
       // If a status for the inerting system changed by operator copy this to the select number and do not read all status values
       IF "DB614_MH_State".InertingMH["DB614_MH_State".ReadDeviceNo].Inert_ON_OFF <> "DB614_MH_State".InertingMH[0].Inert_ON_OFF OR
           "DB614_MH_State".InertingMH["DB614_MH_State".ReadDeviceNo].Enable_Purge <> "DB614_MH_State".InertingMH[0].Enable_Purge
       THEN
           "DB614_MH_State".InertingMH["DB614_MH_State".ReadDeviceNo].Inert_ON_OFF := "DB614_MH_State".InertingMH[0].Inert_ON_OFF;
           "DB614_MH_State".InertingMH["DB614_MH_State".ReadDeviceNo].Enable_Purge := "DB614_MH_State".InertingMH[0].Enable_Purge;
       ELSE
           "DB614_MH_State".InertingMH[0] := "DB614_MH_State".InertingMH["DB614_MH_State".ReadDeviceNo];
       END_IF;

   END_IF;

   // Copy the Status bits after changing
   IF "DB614_MH_State".Write THEN

       "DB614_MH_State".Write := False;

   END_IF;

   // Copy the values if nessesary
   IF "DB704_MH_Value".Write THEN
       "DB604_PV_Mixinghead".Mixinghead["DB614_MH_State".ReadDeviceNo] := "DB604_PV_Mixinghead".Mixinghead[0];
       "DB704_MH_Value".Mixinghead["DB614_MH_State".ReadDeviceNo] := "DB704_MH_Value".Mixinghead[0];
       "DB704_MH_Value".MH_Inerting["DB614_MH_State".ReadDeviceNo] := "DB704_MH_Value".MH_Inerting[0];

       "DB704_MH_Value".Write := False;

   END_IF;

   // Show the actual values every time:
   // 
   "DB604_PV_Mixinghead".Mixinghead[0].Pressure_Connection[1].PV_ActV := "DB604_PV_Mixinghead".Mixinghead["DB614_MH_State".ReadDeviceNo].Pressure_Connection[1].PV_ActV;
   "DB604_PV_Mixinghead".Mixinghead[0].Pressure_Connection[2].PV_ActV := "DB604_PV_Mixinghead".Mixinghead["DB614_MH_State".ReadDeviceNo].Pressure_Connection[2].PV_ActV;
   "DB604_PV_Mixinghead".Mixinghead[0].Pressure_Connection[3].PV_ActV := "DB604_PV_Mixinghead".Mixinghead["DB614_MH_State".ReadDeviceNo].Pressure_Connection[3].PV_ActV;
   "DB604_PV_Mixinghead".Mixinghead[0].Pressure_Connection[4].PV_ActV := "DB604_PV_Mixinghead".Mixinghead["DB614_MH_State".ReadDeviceNo].Pressure_Connection[4].PV_ActV;
   "DB604_PV_Mixinghead".Mixinghead[0].Pressure_Connection[5].PV_ActV := "DB604_PV_Mixinghead".Mixinghead["DB614_MH_State".ReadDeviceNo].Pressure_Connection[5].PV_ActV;
   "DB604_PV_Mixinghead".Mixinghead[0].Pressure_Connection[6].PV_ActV := "DB604_PV_Mixinghead".Mixinghead["DB614_MH_State".ReadDeviceNo].Pressure_Connection[6].PV_ActV;

   "DB604_PV_Mixinghead".Mixinghead[0].Temperature_Connection[1].PV_ActV := "DB604_PV_Mixinghead".Mixinghead["DB614_MH_State".ReadDeviceNo].Temperature_Connection[1].PV_ActV;
   "DB604_PV_Mixinghead".Mixinghead[0].Temperature_Connection[2].PV_ActV := "DB604_PV_Mixinghead".Mixinghead["DB614_MH_State".ReadDeviceNo].Temperature_Connection[2].PV_ActV;
   "DB604_PV_Mixinghead".Mixinghead[0].Temperature_Connection[3].PV_ActV := "DB604_PV_Mixinghead".Mixinghead["DB614_MH_State".ReadDeviceNo].Temperature_Connection[3].PV_ActV;
   "DB604_PV_Mixinghead".Mixinghead[0].Temperature_Connection[4].PV_ActV := "DB604_PV_Mixinghead".Mixinghead["DB614_MH_State".ReadDeviceNo].Temperature_Connection[4].PV_ActV;
   "DB604_PV_Mixinghead".Mixinghead[0].Temperature_Connection[5].PV_ActV := "DB604_PV_Mixinghead".Mixinghead["DB614_MH_State".ReadDeviceNo].Temperature_Connection[5].PV_ActV;
   "DB604_PV_Mixinghead".Mixinghead[0].Temperature_Connection[6].PV_ActV := "DB604_PV_Mixinghead".Mixinghead["DB614_MH_State".ReadDeviceNo].Temperature_Connection[6].PV_ActV;

   "DB604_PV_Mixinghead".Mixinghead[0].SteeringPiston.PV_ActV := "DB604_PV_Mixinghead".Mixinghead["DB614_MH_State".ReadDeviceNo].SteeringPiston.PV_ActV;
   "DB604_PV_Mixinghead".Mixinghead[0].CleaningPiston.PV_ActV := "DB604_PV_Mixinghead".Mixinghead["DB614_MH_State".ReadDeviceNo].CleaningPiston.PV_ActV;
   "DB604_PV_Mixinghead".Mixinghead[0].Inerting.PV_ActV := "DB604_PV_Mixinghead".Mixinghead["DB614_MH_State".ReadDeviceNo].Inerting.PV_ActV;

   // Show the in/ output from MH every time
   "DB123_MH_IO_Signals".MH[0] := "DB123_MH_IO_Signals".MH["DB614_MH_State".ReadDeviceNo];

   // Show the actual information about the selected mixinghead
   "DB614_MH_State".MH_Connection[0] := "DB614_MH_State".MH_Connection["DB614_MH_State".ReadDeviceNo];

   // Information about shot adjustment
   "DB614_MH_State".ShotAdjustMH[0] := "DB614_MH_State".ShotAdjustMH["DB614_MH_State".ReadDeviceNo];
END_FUNCTION

FUNCTION "FC5019_InterfaceInterface" : Void   // FC5019, SCL
{ S7_Optimized_Access := 'FALSE' }
VERSION : 0.1
   VAR_INPUT
      Enable : Bool;
   END_VAR
BEGIN
   // Status: DB612_Hydraulic_State
   // Read all status bits during window is selected and NO button is pressed
     IF "DB119_Interface_Visu".Read THEN
       "DB119_Interface_Visu".MouldCarrer[0] := "DB119_Interface_Visu".MouldCarrer["DB119_Interface_Visu".ReadWriteDeviceNo];
       "DB119_Interface_Visu".APInterface[0] := "DB119_Interface_Visu".APInterface["DB119_Interface_Visu".ReadWriteDeviceNo];
     END_IF;
END_FUNCTION

FUNCTION "FC5020_InterfaceConfig" : Void   // FC5020, SCL
{ S7_Optimized_Access := 'FALSE' }
VERSION : 0.1
   VAR_INPUT
      Enable : Bool;
   END_VAR
BEGIN

   // Values:  "DB1200_ProCanConf" 
     IF "DB1200_ProCanConf".Read OR "DB1200_ProCanConf".Write OR "DB1200_ProCanConf".Copy THEN
       IF "DB1200_ProCanConf".Read THEN
         "DB1200_ProCanConf".ProCanConf[0] := "DB1200_ProCanConf".ProCanConf["DB1200_ProCanConf".ReadWriteDeviceNo];
         "DB1200_ProCanConf".Read := FALSE;
       END_IF;
       IF "DB1200_ProCanConf".Write THEN
         "DB1200_ProCanConf".ProCanConf["DB1200_ProCanConf".ReadWriteDeviceNo] := "DB1200_ProCanConf".ProCanConf[0];
         "DB1200_ProCanConf".Write := FALSE;
       END_IF;
         IF "DB1200_ProCanConf".CopyDeviceNO >0 THEN
         IF "DB1200_ProCanConf".Copy THEN
             "DB1200_ProCanConf".ProCanConf["DB1200_ProCanConf".CopyDeviceNO] := "DB1200_ProCanConf".ProCanConf[0];
             "DB1200_ProCanConf".Copy := FALSE;
             "DB1200_ProCanConf".CopyDeviceNO := 0;
         END_IF;
        END_IF;
      END_IF;    

   // Values:  "DB1232_ProCanIO_MH" 
     IF "DB1232_ProCanIO_MH".Read OR "DB1232_ProCanIO_MH".Write OR "DB1232_ProCanIO_MH".Copy THEN
       IF "DB1232_ProCanIO_MH".Read THEN
         "DB1232_ProCanIO_MH".AddressMH[0] := "DB1232_ProCanIO_MH".AddressMH["DB1232_ProCanIO_MH".ReadWriteDeviceNo];
         "DB1232_ProCanIO_MH".Read := FALSE;
       END_IF;
       IF "DB1232_ProCanIO_MH".Write THEN
         "DB1232_ProCanIO_MH".AddressMH["DB1232_ProCanIO_MH".ReadWriteDeviceNo] := "DB1232_ProCanIO_MH".AddressMH[0];
         "DB1232_ProCanIO_MH".Write := FALSE;
       END_IF;
         IF "DB1232_ProCanIO_MH".CopyDeviceNO >0 THEN
         IF "DB1232_ProCanIO_MH".Copy THEN
             "DB1232_ProCanIO_MH".AddressMH["DB1232_ProCanIO_MH".CopyDeviceNO] := "DB1232_ProCanIO_MH".AddressMH[0];
             "DB1232_ProCanIO_MH".Copy := FALSE;
             "DB1232_ProCanIO_MH".CopyDeviceNO := 0;
         END_IF;
        END_IF;
      END_IF;

   // Values:  "DB1233_ProCanIO_Flow" 
     IF "DB1233_ProCanIO_Flow".Read OR "DB1233_ProCanIO_Flow".Write OR "DB1233_ProCanIO_Flow".Copy THEN
       IF "DB1233_ProCanIO_Flow".Read THEN
         "DB1233_ProCanIO_Flow".AddressFlow[0] := "DB1233_ProCanIO_Flow".AddressFlow["DB1233_ProCanIO_Flow".ReadWriteDeviceNo];
         "DB1233_ProCanIO_Flow".Read := FALSE;
       END_IF;
       IF "DB1233_ProCanIO_Flow".Write THEN
         "DB1233_ProCanIO_Flow".AddressFlow["DB1233_ProCanIO_Flow".ReadWriteDeviceNo] := "DB1233_ProCanIO_Flow".AddressFlow[0];
         "DB1233_ProCanIO_Flow".Write := FALSE;
       END_IF;
         IF "DB1233_ProCanIO_Flow".CopyDeviceNO >0 THEN
         IF "DB1233_ProCanIO_Flow".Copy THEN
             "DB1233_ProCanIO_Flow".AddressFlow["DB1233_ProCanIO_Flow".CopyDeviceNO] := "DB1233_ProCanIO_Flow".AddressFlow[0];
             "DB1233_ProCanIO_Flow".Copy := FALSE;
             "DB1233_ProCanIO_Flow".CopyDeviceNO := 0;
         END_IF;
        END_IF;
      END_IF;
END_FUNCTION

FUNCTION "FC5030_InterfaceactualMHValue" : Void   // FC5030, SCL
{ S7_Optimized_Access := 'FALSE' }
VERSION : 0.1
   VAR_INPUT
      IN_MachineNo : Int;
   END_VAR
   VAR_TEMP
      N : Int;
      i : Int;
      AmountComponent : Int;
      Temp_MachineNo : Byte;
   END_VAR
BEGIN
   // Baustein zur Ermittlung der akteullen Mischkopf- Informationen
   // 
   // 1. Maschine ist im Ruhestand, Kein Kreislauf oder Zyxklus aktiv
   //    Die Werte des zuerst freigegebenen Mischkopfes an dieser Maschine werden angezeigt
   //  
   #Temp_MachineNo := INT_TO_BYTE(#IN_MachineNo);
   //  
   "DB619_State_MPart".ActMHInerting[#IN_MachineNo].Total_Flow_N2_Visu := "DB614_MH_State".InertingMH[1].Total_Flow_N2_Visu;

   IF NOT "DB619_State_MPart".Recirculation[#IN_MachineNo].Is_active AND
      NOT "DB619_State_MPart".Cycle[#IN_MachineNo].running THEN

      "DB619_State_MPart".ActMHComponent[1].OP_Manual := 0;
      "DB619_State_MPart".ActMHComponent[1].OP_Automatic := 0;
      "DB619_State_MPart".ActMHComponent[1].OP_Service := 0;

     FOR #N := 1 TO "DB790_PlantParameter".AmountMH DO

       IF "DB704_MH_Value".Mixinghead[#N].MH_Active AND
           "DB704_MH_Value".Mixinghead[#N].MachineNumber = #Temp_MachineNo THEN

         "DB619_State_MPart".ActMHPressureMa[#IN_MachineNo].Comp[1] :=  "DB604_PV_Mixinghead".Mixinghead[#N].Pressure_Connection[1].PV_ActV.Value;
         "DB619_State_MPart".ActMHPressureMa[#IN_MachineNo].Comp[2] :=  "DB604_PV_Mixinghead".Mixinghead[#N].Pressure_Connection[2].PV_ActV.Value;
         "DB619_State_MPart".ActMHPressureMa[#IN_MachineNo].Comp[3] :=  "DB604_PV_Mixinghead".Mixinghead[#N].Pressure_Connection[3].PV_ActV.Value;
         "DB619_State_MPart".ActMHPressureMa[#IN_MachineNo].Comp[4] :=  "DB604_PV_Mixinghead".Mixinghead[#N].Pressure_Connection[4].PV_ActV.Value;
         "DB619_State_MPart".ActMHPressureMa[#IN_MachineNo].Comp[5] :=  "DB604_PV_Mixinghead".Mixinghead[#N].Pressure_Connection[5].PV_ActV.Value;
         "DB619_State_MPart".ActMHPressureMa[#IN_MachineNo].Comp[6] :=  "DB604_PV_Mixinghead".Mixinghead[#N].Pressure_Connection[6].PV_ActV.Value;
         "DB619_State_MPart".ActMHTemperatureMa[#IN_MachineNo].Comp[1] :=  "DB604_PV_Mixinghead".Mixinghead[#N].Temperature_Connection[1].PV_ActV.Value;
         "DB619_State_MPart".ActMHTemperatureMa[#IN_MachineNo].Comp[2] :=  "DB604_PV_Mixinghead".Mixinghead[#N].Temperature_Connection[2].PV_ActV.Value;
         "DB619_State_MPart".ActMHTemperatureMa[#IN_MachineNo].Comp[3] :=  "DB604_PV_Mixinghead".Mixinghead[#N].Temperature_Connection[3].PV_ActV.Value;
         "DB619_State_MPart".ActMHTemperatureMa[#IN_MachineNo].Comp[4] :=  "DB604_PV_Mixinghead".Mixinghead[#N].Temperature_Connection[4].PV_ActV.Value;
         "DB619_State_MPart".ActMHTemperatureMa[#IN_MachineNo].Comp[5] :=  "DB604_PV_Mixinghead".Mixinghead[#N].Temperature_Connection[5].PV_ActV.Value;
         "DB619_State_MPart".ActMHTemperatureMa[#IN_MachineNo].Comp[6] :=  "DB604_PV_Mixinghead".Mixinghead[#N].Temperature_Connection[6].PV_ActV.Value;

         "DB619_State_MPart".ActMHComponent[#IN_MachineNo].No := "DB704_MH_Value".Mixinghead[#N].#AmountComponent;
         "DB619_State_MPart".ActMHComponent[#IN_MachineNo].Name[1] := "DB614_MH_State".MH_Connection[#N].Name[1];
         "DB619_State_MPart".ActMHComponent[#IN_MachineNo].Name[2] := "DB614_MH_State".MH_Connection[#N].Name[2];
         "DB619_State_MPart".ActMHComponent[#IN_MachineNo].Name[3] := "DB614_MH_State".MH_Connection[#N].Name[3];
         "DB619_State_MPart".ActMHComponent[#IN_MachineNo].Name[4] := "DB614_MH_State".MH_Connection[#N].Name[4];
         "DB619_State_MPart".ActMHComponent[#IN_MachineNo].Name[5] := "DB614_MH_State".MH_Connection[#N].Name[5];
         "DB619_State_MPart".ActMHComponent[#IN_MachineNo].Name[6] := "DB614_MH_State".MH_Connection[#N].Name[6];
         "DB619_State_MPart".ActMHComponent[#IN_MachineNo].colour[1]:= "DB614_MH_State".MH_Connection[#N].colour[1];
         "DB619_State_MPart".ActMHComponent[#IN_MachineNo].colour[2] := "DB614_MH_State".MH_Connection[#N].colour[2];
         "DB619_State_MPart".ActMHComponent[#IN_MachineNo].colour[3] := "DB614_MH_State".MH_Connection[#N].colour[3];
         "DB619_State_MPart".ActMHComponent[#IN_MachineNo].colour[4] := "DB614_MH_State".MH_Connection[#N].colour[4];
         "DB619_State_MPart".ActMHComponent[#IN_MachineNo].colour[5] := "DB614_MH_State".MH_Connection[#N].colour[5];
         "DB619_State_MPart".ActMHComponent[#IN_MachineNo].colour[6] := "DB614_MH_State".MH_Connection[#N].colour[6];


         RETURN;
       END_IF;
     END_FOR;
   END_IF;
   // 
   // 2. Beim Kreislauf oder Zyklus werden die Werte der aktuellen USE angezeigt
   //    Diese Werte werden auch für die Schussprotokollierung verwendet!
   //    Wenn kein Kreislauf dann "0"

   #N := "DB619_State_MPart".SWU[#IN_MachineNo].ActualSWU;

   "DB619_State_MPart".ActMHComponent[1].OP_Manual := "DB123_MH_IO_Signals".MH[#N].IN.MH_Manual_Mode;
   "DB619_State_MPart".ActMHComponent[1].OP_Automatic := "DB123_MH_IO_Signals".MH[#N].IN.MH_Auto_Mode;
   "DB619_State_MPart".ActMHComponent[1].OP_Service := NOT "DB614_MH_State".MH_Status[#N].Switch_Service_ON_OFF OR
   ("DB619_State_MPart".Operationmode[1].Operation AND "DB619_State_MPart".ShotMa[1].ShotData.ShotDisabled AND "DB619_State_MPart".Operationmode[1].Auto AND NOT "DB619_State_MPart".Operationmode[1].Test);

   // IF "DB123_MH_IO_Signals".MH[#N].OUT.MH.ServiceProduction = 0 THEN
   //     "DB619_State_MPart".ActMHComponent[1].OP_Service := 1;
   // END_IF;


   "DB619_State_MPart".ActMHPressureMa[#IN_MachineNo].Comp[1] := "DB604_PV_Mixinghead".Mixinghead[#N].Pressure_Connection[1].PV_ActV.Value;
   "DB619_State_MPart".ActMHPressureMa[#IN_MachineNo].Comp[2] := "DB604_PV_Mixinghead".Mixinghead[#N].Pressure_Connection[2].PV_ActV.Value;
   "DB619_State_MPart".ActMHPressureMa[#IN_MachineNo].Comp[3] := "DB604_PV_Mixinghead".Mixinghead[#N].Pressure_Connection[3].PV_ActV.Value;
   "DB619_State_MPart".ActMHPressureMa[#IN_MachineNo].Comp[4] := "DB604_PV_Mixinghead".Mixinghead[#N].Pressure_Connection[4].PV_ActV.Value;
   "DB619_State_MPart".ActMHPressureMa[#IN_MachineNo].Comp[5] := "DB604_PV_Mixinghead".Mixinghead[#N].Pressure_Connection[5].PV_ActV.Value;
   "DB619_State_MPart".ActMHPressureMa[#IN_MachineNo].Comp[6] := "DB604_PV_Mixinghead".Mixinghead[#N].Pressure_Connection[6].PV_ActV.Value;
   "DB619_State_MPart".ActMHTemperatureMa[#IN_MachineNo].Comp[1] := "DB604_PV_Mixinghead".Mixinghead[#N].Temperature_Connection[1].PV_ActV.Value;
   "DB619_State_MPart".ActMHTemperatureMa[#IN_MachineNo].Comp[2] := "DB604_PV_Mixinghead".Mixinghead[#N].Temperature_Connection[2].PV_ActV.Value;
   "DB619_State_MPart".ActMHTemperatureMa[#IN_MachineNo].Comp[3] := "DB604_PV_Mixinghead".Mixinghead[#N].Temperature_Connection[3].PV_ActV.Value;
   "DB619_State_MPart".ActMHTemperatureMa[#IN_MachineNo].Comp[4] := "DB604_PV_Mixinghead".Mixinghead[#N].Temperature_Connection[4].PV_ActV.Value;
   "DB619_State_MPart".ActMHTemperatureMa[#IN_MachineNo].Comp[5] := "DB604_PV_Mixinghead".Mixinghead[#N].Temperature_Connection[5].PV_ActV.Value;
   "DB619_State_MPart".ActMHTemperatureMa[#IN_MachineNo].Comp[6] := "DB604_PV_Mixinghead".Mixinghead[#N].Temperature_Connection[6].PV_ActV.Value;

   "DB619_State_MPart".ActMHComponent[#IN_MachineNo].No := "DB704_MH_Value".Mixinghead[#N].#AmountComponent;
   "DB619_State_MPart".ActMHComponent[#IN_MachineNo].Name[1] := "DB614_MH_State".MH_Connection[#N].Name[1];
   "DB619_State_MPart".ActMHComponent[#IN_MachineNo].Name[2] := "DB614_MH_State".MH_Connection[#N].Name[2];
   "DB619_State_MPart".ActMHComponent[#IN_MachineNo].Name[3] := "DB614_MH_State".MH_Connection[#N].Name[3];
   "DB619_State_MPart".ActMHComponent[#IN_MachineNo].Name[4] := "DB614_MH_State".MH_Connection[#N].Name[4];
   "DB619_State_MPart".ActMHComponent[#IN_MachineNo].Name[5] := "DB614_MH_State".MH_Connection[#N].Name[5];
   "DB619_State_MPart".ActMHComponent[#IN_MachineNo].Name[6] := "DB614_MH_State".MH_Connection[#N].Name[6];
   "DB619_State_MPart".ActMHComponent[#IN_MachineNo].colour[1] := "DB614_MH_State".MH_Connection[#N].colour[1];
   "DB619_State_MPart".ActMHComponent[#IN_MachineNo].colour[2] := "DB614_MH_State".MH_Connection[#N].colour[2];
   "DB619_State_MPart".ActMHComponent[#IN_MachineNo].colour[3] := "DB614_MH_State".MH_Connection[#N].colour[3];
   "DB619_State_MPart".ActMHComponent[#IN_MachineNo].colour[4] := "DB614_MH_State".MH_Connection[#N].colour[4];
   "DB619_State_MPart".ActMHComponent[#IN_MachineNo].colour[5] := "DB614_MH_State".MH_Connection[#N].colour[5];
   "DB619_State_MPart".ActMHComponent[#IN_MachineNo].colour[6] := "DB614_MH_State".MH_Connection[#N].colour[6];

   // 3. Einige Werte werden dann nur für die Schussprotokollierung verwendet:
   // 
   //  #N := "DB619_State_MPart".SWU[#IN_MachineNo].ActualSWU;
     // Tanktemperatur:
   //  "DB919_ShotResultMach".ShotResult_Ma[#IN_MachineNo].Component.Comp[1].Temperature := "DB602_PV_Tank".Tank[1].Temp.PV_ActV.Value;
   //
   //
END_FUNCTION

FUNCTION "FC5031_InterfaceMachineGeneral" : Void   // FC5031, SCL
{ S7_Optimized_Access := 'FALSE' }
VERSION : 0.1
BEGIN
   // Status: DB619_State_MPart
   // Values: DB700_Machine
   // Faults: DB829_Error_Machine
   // 
   // Read the Values only once after open the window or change the Number
   // 
     IF ("DB619_State_MPart".ReadDeviceNo <> "DB619_State_MPart".ActualDeviceNo) OR "DB619_State_MPart".Read THEN
         "DB619_State_MPart".ActualDeviceNo := "DB619_State_MPart".ReadDeviceNo;

         // Status
         // Setvalues 
         "DB700_Machine".Machine[0] := "DB700_Machine".Machine["DB619_State_MPart".ReadDeviceNo];

         "DB619_State_MPart".Read := FALSE;

     END_IF;

     IF "DB619_State_MPart".Write THEN
         // Set the Button to the right destination
         // Values 
         "DB700_Machine".Machine["DB619_State_MPart".ReadDeviceNo] := "DB700_Machine".Machine[0];
         // Reset write signal
     END_IF;

     "DB619_State_MPart".Write := FALSE;
END_FUNCTION

FUNCTION "FC5032_Last10Shot" : Void   // FC5032, SCL
{ S7_Optimized_Access := 'FALSE' }
VERSION : 0.1
   VAR_INPUT
      IN_MachineNo : Int;
   END_VAR
   VAR_TEMP
      N : Int;
   END_VAR
BEGIN
     IF "DB918_ShotResultlast10".NewData THEN
     FOR #N := 1 TO 19 DO
       "DB918_ShotResultlast10".RealShot[21-#N] := "DB918_ShotResultlast10".RealShot[20-#N];
     END_FOR;

   //  "DB918_ShotResultlast10".RealShot[1].PartNo :=
     "DB918_ShotResultlast10".RealShot[1].PartNo :=  "DB919_ShotResultMach".ShotResult_Ma[#IN_MachineNo].General.ShotNo;
     "DB918_ShotResultlast10".RealShot[1].PartCounter :=  "DB919_ShotResultMach".ShotResult_Ma[#IN_MachineNo].General.PartID;
     "DB918_ShotResultlast10".RealShot[1].MHNo := "DB919_ShotResultMach".ShotResult_Ma[#IN_MachineNo].General.MH_No;
     "DB918_ShotResultlast10".RealShot[1].FoamingTime := "DB919_ShotResultMach".ShotResult_Ma[#IN_MachineNo].General.FoamingTime;
     "DB918_ShotResultlast10".RealShot[1].PartWeight := "DB919_ShotResultMach".ShotResult_Ma[#IN_MachineNo].General.PartWeight;
     "DB918_ShotResultlast10".RealShot[1].StationNo := "DB919_ShotResultMach".ShotResult_Ma[#IN_MachineNo].General.StationNo;
     "DB918_ShotResultlast10".RealShot[1].Machine_No := "DB919_ShotResultMach".ShotResult_Ma[#IN_MachineNo].General.Machine_No;
     "DB918_ShotResultlast10".RealShot[1].Nitrogen := "DB919_ShotResultMach".ShotResult_Ma[#IN_MachineNo].General.NitrogenValue_Inerting;

     FOR #N := 1 TO 6 DO
       "DB918_ShotResultlast10".RealShot[1].Name[#N] := "DB919_ShotResultMach".ShotResult_Ma[#IN_MachineNo].Component.Comp[#N].Name;
       "DB918_ShotResultlast10".RealShot[1].Flow[#N] := "DB919_ShotResultMach".ShotResult_Ma[#IN_MachineNo].Component.Comp[#N].Flow;
       "DB918_ShotResultlast10".RealShot[1].Pressure[#N] := "DB919_ShotResultMach".ShotResult_Ma[#IN_MachineNo].Component.Comp[#N].PressureMH;
       "DB918_ShotResultlast10".RealShot[1].Temperature[#N] := "DB919_ShotResultMach".ShotResult_Ma[#IN_MachineNo].Component.Comp[#N].TemperatureMH;
       "DB918_ShotResultlast10".RealShot[1].MaterialConsumption[#N] := "DB919_ShotResultMach".ShotResult_Ma[#IN_MachineNo].Component.Comp[#N].MaterialConsumption;
       "DB918_ShotResultlast10".RealShot[1].Mixingratio[#N] :=  "DB919_ShotResultMach".ShotResult_Ma[#IN_MachineNo].Component.Comp[#N].Mixingratio;
   //  "DB918_ShotResultlast10".RealShot[1].StausBitWarning :=
     END_FOR;


   //  "DB918_ShotResultlast10".RealShot[1].PartShotDisableService :=
     "DB918_ShotResultlast10".RealShot[1].StatusBitFaultGroup1 := "DB919_ShotResultMach".ShotResult_Ma[#IN_MachineNo].General.ShotState[0];
     "DB918_ShotResultlast10".RealShot[1].StatusBitStopCycleDuringShot := "DB919_ShotResultMach".ShotResult_Ma[#IN_MachineNo].General.ShotState[1];
     "DB918_ShotResultlast10".RealShot[1].PartShotDisableService :="DB919_ShotResultMach".ShotResult_Ma[#IN_MachineNo].General.ShotState[2];
     "DB918_ShotResultlast10".RealShot[1].StatusBitManualShot :="DB919_ShotResultMach".ShotResult_Ma[#IN_MachineNo].General.ShotState[3];
     "DB918_ShotResultlast10".RealShot[1].StatusBitAutomaticShot := NOT "DB919_ShotResultMach".ShotResult_Ma[#IN_MachineNo].General.ShotState[3];

   //  "DB918_ShotResultlast10".RealShot[1].StatusBitWarningFlow :=
   //  "DB918_ShotResultlast10".RealShot[1].StatusBitAlarmFlow :=
   //  "DB918_ShotResultlast10".RealShot[1].StatusBitWarningWeight :=
   //  "DB918_ShotResultlast10".RealShot[1].StatusBitAlarmWeight :=
   //  "DB918_ShotResultlast10".RealShot[1].StatusBitWarningFoamingTime :=
   //  "DB918_ShotResultlast10".RealShot[1].StatusBitAlarmFoamingTime :=


   // Möglicher Filter einbauen!
     FOR #N := 1 TO 10 DO
       "DB918_ShotResultlast10".FilteredShot[#N] := "DB918_ShotResultlast10".RealShot[#N];
     END_FOR;




     "DB918_ShotResultlast10".NewData := 0;
   END_IF;
END_FUNCTION

FUNCTION "FC5900_InterfaceRobots" : Void   // FC5900, SCL
{ S7_Optimized_Access := 'FALSE' }
VERSION : 0.1
   VAR_INPUT
      Enable : Bool;
   END_VAR
BEGIN
   // Status: DB1901_Config_Robots 
   // Read all status bits during window is selected and NO button is pressed
   IF "DB1901_Config_Robots".Read AND NOT "DB1901_Config_Robots".Write THEN
       "DB1901_Config_Robots".Config_Robots[0] := "DB1901_Config_Robots".Config_Robots["DB1900_IF_Robots".ReadWriteDeviceNo];
   END_IF;
   // Set the Button to the right destination
   IF "DB1901_Config_Robots".Read AND "DB1901_Config_Robots".Write THEN
       "DB1901_Config_Robots".Config_Robots["DB1900_IF_Robots".ReadWriteDeviceNo] := "DB1901_Config_Robots".Config_Robots[0];
       "DB1901_Config_Robots".Write := False;
   END_IF;

   // Status: DB1900_IF_Robots 
   // Read all status bits during window is selected and NO button is pressed
   IF "DB1900_IF_Robots".Read AND NOT "DB1900_IF_Robots".Write THEN
       "DB1900_IF_Robots".Switch_Robots[0] := "DB1900_IF_Robots".Switch_Robots["DB1900_IF_Robots".ReadWriteDeviceNo];
       "DB1900_IF_Robots".State_Robots[0] := "DB1900_IF_Robots".State_Robots["DB1900_IF_Robots".ReadWriteDeviceNo];
       "DB1900_IF_Robots".Faults_Robots[0] := "DB1900_IF_Robots".Faults_Robots["DB1900_IF_Robots".ReadWriteDeviceNo];
   END_IF;
   // Set the Button to the right destination
   IF "DB1900_IF_Robots".Read AND "DB1900_IF_Robots".Write THEN
       "DB1900_IF_Robots".Switch_Robots["DB1900_IF_Robots".ReadWriteDeviceNo] := "DB1900_IF_Robots".Switch_Robots[0];
       "DB1900_IF_Robots".Write := False;
   END_IF;
END_FUNCTION

FUNCTION "FC5901_generalFunction" : Void   // FC5901, SCL
{ S7_Optimized_Access := 'FALSE' }
VERSION : 0.1
   VAR_OUTPUT
      StartCycle : Bool;
      EnableMCatPos1 : Bool;
      TestShotActiv : Bool;
      AtPos1or2 : Bool;
   END_VAR
   VAR_TEMP
      Interface : Int;
      Temp_StartCycle : Bool;
      Temp_EnableMCatPos1 : Bool;
      Temp_TestShotActiv : Bool;
      Temp_AtPos1or2 : Bool;
   END_VAR
BEGIN
   // create general signals for the interface between robots and machine
   // 
   #Temp_StartCycle := 0;
   FOR #Interface := 1 TO "DB790_PlantParameter".AmountMouldCarrier DO
       IF #Interface >16 THEN
           EXIT;
       ELSIF "DB1901_Config_Robots".Config_Robots[1].ForInterface[#Interface] = True AND #Interface <=16  THEN
           #Temp_StartCycle := #Temp_StartCycle OR "DB110_Interf_Program_M1".Status_IF[#Interface].Start_to_Cycle;
       END_IF;
   END_FOR;
   #StartCycle := #Temp_StartCycle;

   //------------------------------
   //
   #Temp_EnableMCatPos1 := 0;
   FOR #Interface := 1 TO "DB790_PlantParameter".AmountMouldCarrier DO
       IF #Interface >16 THEN
           EXIT;
       ELSIF "DB1901_Config_Robots".Config_Robots[1].ForInterface[#Interface] = True AND #Interface <=16 THEN
           #Temp_EnableMCatPos1 := #Temp_EnableMCatPos1 OR ("DB005_RS<->Extern".MC_Interface[#Interface].Data_from_MC.Shot_release AND "DB110_Interf_Program_M1".Status_IF[#Interface].IF_is_on_1_Position);
       END_IF;
   END_FOR;
   #EnableMCatPos1 := #Temp_EnableMCatPos1;

   //------------------------------
   //
   #Temp_TestShotActiv := 0;
   IF "DB110_Interf_Program_M1".FIRST = BYTE_TO_INT("DB1901_Config_Robots".Config_Robots[1].InterfaceForTestShot) THEN
       #Temp_TestShotActiv := TRUE;
   END_IF;
   #TestShotActiv := #Temp_TestShotActiv;

   //------------------------------
   //
   #Temp_AtPos1or2 := 0;
   FOR #Interface := 1 TO "DB790_PlantParameter".AmountMouldCarrier DO
       IF #Interface >16 THEN
           EXIT;
       ELSIF "DB1901_Config_Robots".Config_Robots[1].ForInterface[#Interface] = True AND #Interface <=16 THEN
           #Temp_AtPos1or2 := #Temp_AtPos1or2 OR "DB110_Interf_Program_M1".Status_IF[#Interface].IF_is_on_1_Position OR  "DB110_Interf_Program_M1".Status_IF[#Interface].IF_is_on_2_Position;
       END_IF;
   END_FOR;
   #AtPos1or2 := #Temp_AtPos1or2;

   //------------------------------
   //
   "DB614_MH_State".MH_Status[BYTE_TO_INT("DB1901_Config_Robots".Config_Robots[1].MHNumber)].OpenMHEnableExtern := #EnableMCatPos1;
END_FUNCTION

FUNCTION "FC_ActPressureMeteringUnit" : Void   // FC7001, SCL
{ S7_Optimized_Access := 'FALSE' }
VERSION : 0.1
   VAR_TEMP
      DInt_dummy : Real;
      N : Int;
   END_VAR
BEGIN

   FOR #N := 1 TO "DB790_PlantParameter".AmountMeteringUnits DO
       "FC920_PV_Calc_Act_Value"(IN_Act_Value_read := TRUE,
                                 IN_Act_Value_ext := FALSE,
                                 IN_Ext_Value := #DInt_dummy,
                                 IN_Read_Double := FALSE,
                                 IN_FLT_Needful := TRUE,
                                 IN_FLT_Reset := "DB009_Faults".Faults_Reset_FKT_M1,
                                 IO_Any_ArrayPV := "DB608_PV_Metering".Metering[#N].Pressure,
                                 IO_Fault_Sensor := "DB823_Error_Metering".Pressure_Component[#N].Sensor_FLT_broken_wire,
                                 IO_New_Fault := "DB009_Faults".Faultschanging_M1,
                                 IO_FLT_Level_3 := "DB009_Faults".Faults_FKT_Grp_3_M1);

       "FC920_PV_Calc_Act_Value"(IN_Act_Value_read := "DB613_Komponent_State".MeteringPump[#N].Selection_Feedingpump,
                                 IN_Act_Value_ext := FALSE,
                                 IN_Ext_Value := #DInt_dummy,
                                 IN_Read_Double := FALSE,
                                 IN_FLT_Needful := TRUE,
                                 IN_FLT_Reset := "DB009_Faults".Faults_Reset_FKT_M1,
                                 IO_Any_ArrayPV := "DB608_PV_Metering".Metering[#N].Pre_Pressure,
                                 IO_Fault_Sensor := "DB823_Error_Metering".PrePressure_Component[#N].Sensor_FLT_broken_wire,
                                 IO_New_Fault := "DB009_Faults".Faultschanging_M1,
                                 IO_FLT_Level_3 := "DB009_Faults".Faults_FKT_Grp_3_M1);

       ;
   END_FOR;
END_FUNCTION

FUNCTION "FC_ActValueMH" : Void   // FC7002, SCL
{ S7_Optimized_Access := 'FALSE' }
VERSION : 0.1
   VAR_TEMP
      MHNumber : Int;
      MHConnection : Int;
      DInt_dummy : Real;
      Temp_ConMHConnected : Bool;
      Temp_WithInerting : Bool;
      Temp_WithAnaCP : Bool;
      Temp_WithAnaMH : Bool;
   END_VAR
BEGIN

   #MHNumber := 1;
   #MHConnection := 1;

   FOR #MHNumber := 1 TO "DB790_PlantParameter".AmountMH DO

       FOR #MHConnection := 1 TO BYTE_TO_INT("DB704_MH_Value".Mixinghead[#MHNumber].AmountComponent) DO
           #Temp_ConMHConnected := ("DB704_MH_Value".Mixinghead[#MHNumber].MH_Connection[#MHConnection].Pump_No > 0 ) AND "PN_AI".Module[#MHNumber+1].AI8.Active;

           // Temperature at the mixinghead connection
           "FC920_PV_Calc_Act_Value"(IN_Act_Value_read:=#Temp_ConMHConnected,
                                     IN_Act_Value_ext:=FALSE,
                                     IN_Ext_Value:=#DInt_dummy,
                                     IN_Read_Double:=FALSE,
                                     IN_FLT_Needful:=TRUE,
                                     IN_FLT_Reset:="DB009_Faults".Faults_Reset_FKT_M1,
                                     IO_Any_ArrayPV:="DB604_PV_Mixinghead".Mixinghead[#MHNumber].Temperature_Connection[#MHConnection],
                                     IO_Fault_Sensor:="DB824_Error_MH_CP".Temperature[#MHConnection, #MHNumber].Sensor_FLT_broken_wire,
                                     IO_New_Fault:="DB009_Faults".Faultschanging_M1,
                                     IO_FLT_Level_3:="DB009_Faults".Faults_FKT_Grp_3_M1);

           // Pressure at the mixinghead connection
           "FC920_PV_Calc_Act_Value"(IN_Act_Value_read := #Temp_ConMHConnected,
                                     IN_Act_Value_ext := FALSE,
                                     IN_Ext_Value := #DInt_dummy,
                                     IN_Read_Double := FALSE,
                                     IN_FLT_Needful := TRUE,
                                     IN_FLT_Reset := "DB009_Faults".Faults_Reset_FKT_M1,
                                     IO_Any_ArrayPV := "DB604_PV_Mixinghead".Mixinghead[#MHNumber].Pressure_Connection[#MHConnection],
                                     IO_Fault_Sensor := "DB824_Error_MH_CP".Pressure[#MHConnection, #MHNumber].Sensor_FLT_broken_wire,
                                     IO_New_Fault := "DB009_Faults".Faultschanging_M1,
                                     IO_FLT_Level_3 := "DB009_Faults".Faults_FKT_Grp_3_M1);

       END_FOR;

       // Inerting Flow at the mixinghead connection
       #Temp_WithInerting := "DB1232_ProCanIO_MH".AddressMH[#MHNumber].Ref_OK AND "DB704_MH_Value".Mixinghead[#MHNumber].WithInerting;
       "FC920_PV_Calc_Act_Value"(IN_Act_Value_read := #Temp_WithInerting,
                                 IN_Act_Value_ext := FALSE,
                                 IN_Ext_Value := #DInt_dummy,
                                 IN_Read_Double := FALSE,
                                 IN_FLT_Needful := TRUE,
                                 IN_FLT_Reset := "DB009_Faults".Faults_Reset_FKT_M1,
                                 IO_Any_ArrayPV := "DB604_PV_Mixinghead".Mixinghead[#MHNumber].Inerting,
                                 IO_Fault_Sensor := "DB824_Error_MH_CP".InertingBlowOut_MH[#MHNumber].Sensor_FLT_broken_wire,
                                 IO_New_Fault := "DB009_Faults".Faultschanging_M1,
                                 IO_FLT_Level_3 := "DB009_Faults".Faults_FKT_Grp_3_M1);

       // position of analouge cleaning pisteon
       #Temp_WithAnaCP :=
       ("DB704_MH_Value".Mixinghead[#MHNumber].Cleaning_Piston.StepCleaningPiston OR
       "DB704_MH_Value".Mixinghead[#MHNumber].Cleaning_Piston.ContrCleaningPiston) AND
       "DB1232_ProCanIO_MH".AddressMH[#MHNumber].Ref_OK;
       "FC920_PV_Calc_Act_Value"(IN_Act_Value_read := #Temp_WithAnaCP,
                                 IN_Act_Value_ext := FALSE,
                                 IN_Ext_Value := #DInt_dummy,
                                 IN_Read_Double := FALSE,
                                 IN_FLT_Needful := TRUE,
                                 IN_FLT_Reset := "DB009_Faults".Faults_Reset_FKT_M1,
                                 IO_Any_ArrayPV := "DB604_PV_Mixinghead".Mixinghead[#MHNumber].CleaningPiston,
                                 IO_Fault_Sensor := "DB824_Error_MH_CP".CleaningPiston[#MHNumber].Sensor_FLT_broken_wire,
                                 IO_New_Fault := "DB009_Faults".Faultschanging_M1,
                                 IO_FLT_Level_3 := "DB009_Faults".Faults_FKT_Grp_3_M1);

       "DB614_MH_State".InertingMH[#MHNumber].Actual_Flow_N2 := "DB604_PV_Mixinghead".Mixinghead[#MHNumber].Inerting.PV_ActV.Value;

       // position of analouge mixinghead
       #Temp_WithAnaMH := "DB704_MH_Value".Mixinghead[#MHNumber].Conf_MHControled AND "DB1232_ProCanIO_MH".AddressMH[#MHNumber].Ref_OK;
       "FC920_PV_Calc_Act_Value"(IN_Act_Value_read := #Temp_WithAnaMH,
                                 IN_Act_Value_ext := FALSE,
                                 IN_Ext_Value := #DInt_dummy,
                                 IN_Read_Double := FALSE,
                                 IN_FLT_Needful := TRUE,
                                 IN_FLT_Reset := "DB009_Faults".Faults_Reset_FKT_M1,
                                 IO_Any_ArrayPV := "DB604_PV_Mixinghead".Mixinghead[#MHNumber].SteeringPiston,
                                 IO_Fault_Sensor := "DB824_Error_MH_CP".SteeringPiston[#MHNumber].Sensor_FLT_broken_wire,
                                 IO_New_Fault := "DB009_Faults".Faultschanging_M1,
                                 IO_FLT_Level_3 := "DB009_Faults".Faults_FKT_Grp_3_M1);

   END_FOR;
END_FUNCTION

FUNCTION "FC_ToleranceValuesMH" : Void   // FC7003, SCL
{ S7_Optimized_Access := 'FALSE' }
VERSION : 0.1
   VAR_INPUT
      CompForShot : Array[1..16] of Bool;
      SwitchOffControl : Bool;
   END_VAR
   VAR_TEMP
      MHNumber : Int;
      MHConnection : Int;
      TempUSEOpen : Array[1..16] of Bool;
      TempStartTolTest : Bool;
      TempEnableTolTestPressure : Bool;
      EnableTolTestPressure : Bool;
   END_VAR
BEGIN

   #MHNumber := 1;
   #MHConnection := 1;

   #TempUSEOpen[1] := "DB619_State_MPart".SWU[1].Open_SWU_allone."01";
   #TempUSEOpen[2] := "DB619_State_MPart".SWU[1].Open_SWU_allone."02";
   #TempUSEOpen[3] := "DB619_State_MPart".SWU[1].Open_SWU_allone."03";
   #TempUSEOpen[4] := "DB619_State_MPart".SWU[1].Open_SWU_allone."04";
   #TempUSEOpen[5] := "DB619_State_MPart".SWU[1].Open_SWU_allone."05";
   #TempUSEOpen[6] := "DB619_State_MPart".SWU[1].Open_SWU_allone."06";
   #TempUSEOpen[7] := "DB619_State_MPart".SWU[1].Open_SWU_allone."07";
   #TempUSEOpen[8] := "DB619_State_MPart".SWU[1].Open_SWU_allone."08";
   #TempUSEOpen[9] := "DB619_State_MPart".SWU[1].Open_SWU_allone."09";
   #TempUSEOpen[10] := "DB619_State_MPart".SWU[1].Open_SWU_allone."10";
   #TempUSEOpen[11] := "DB619_State_MPart".SWU[1].Open_SWU_allone."11";
   #TempUSEOpen[12] := "DB619_State_MPart".SWU[1].Open_SWU_allone."12";
   #TempUSEOpen[13] := "DB619_State_MPart".SWU[1].Open_SWU_allone."13";
   #TempUSEOpen[14] := "DB619_State_MPart".SWU[1].Open_SWU_allone."14";
   #TempUSEOpen[15] := "DB619_State_MPart".SWU[1].Open_SWU_allone."15";
   #TempUSEOpen[16] := "DB619_State_MPart".SWU[1].Open_SWU_allone."16";


   FOR #MHNumber := 1 TO "DB790_PlantParameter".AmountMH DO

       FOR #MHConnection := 1 TO BYTE_TO_INT("DB704_MH_Value".Mixinghead[#MHNumber].AmountComponent) DO

           IF "DB704_MH_Value".Mixinghead[#MHNumber].MH_Connection[#MHConnection].Pump_No <> 0 THEN

               IF "DB604_PV_Mixinghead".Mixinghead[#MHNumber].Pressure_Connection[#MHConnection].PV_SetV.Value > 0 THEN
                   #TempEnableTolTestPressure := 1;
               END_IF;

               #TempStartTolTest :=
               #CompForShot["DB704_MH_Value".Mixinghead[#MHNumber].MH_Connection[#MHConnection].Pump_No]
               AND #TempUSEOpen[#MHNumber]
               AND "DB619_State_MPart".Cycle[1].Shotrelease
               AND NOT #SwitchOffControl;

               #EnableTolTestPressure := #TempStartTolTest AND #TempEnableTolTestPressure;

               "FC916_PV_Limits"(IN_Tolerance_Test := #TempStartTolTest,
                                 IN_Reset_Fault := "DB009_Faults".Faults_Reset_FKT_M1,
                                 IO_Any_ArrayPV := "DB604_PV_Mixinghead".Mixinghead[#MHNumber].Temperature_Connection[#MHConnection],
                                 IO_Fault_Warn_upperL := "DB824_Error_MH_CP".Temperature[#MHConnection, #MHNumber].Warning_limit_plus,
                                 IO_Fault_Warn_lowerL := "DB824_Error_MH_CP".Temperature[#MHConnection, #MHNumber].Warning_limit_minus,
                                 IO_Fault_Alarm_upperL := "DB824_Error_MH_CP".Temperature[#MHConnection, #MHNumber].Alarm_limit_plus,
                                 IO_Fault_Alarm_lowerL := "DB824_Error_MH_CP".Temperature[#MHConnection, #MHNumber].Alarm_limit_minus,
                                 IO_New_Fault := "DB009_Faults".Faultschanging_M1,
                                 IO_Fault_Level_1 := "DB009_Faults".Faults_FKT_Grp_1_M1,
                                 IO_Fault_Level_2 := "DB009_Faults".Faults_FKT_Grp_2_M1,
                                 IO_Fault_Level_3 := "DB009_Faults".Faults_FKT_Grp_3_M1);

               "FC916_PV_Limits"(IN_Tolerance_Test := #EnableTolTestPressure,
                                 IN_Reset_Fault := "DB009_Faults".Faults_Reset_FKT_M1,
                                 IO_Any_ArrayPV := "DB604_PV_Mixinghead".Mixinghead[#MHNumber].Pressure_Connection[#MHConnection],
                                 IO_Fault_Warn_upperL := "DB824_Error_MH_CP".Pressure[#MHConnection, #MHNumber].Warning_limit_plus,
                                 IO_Fault_Warn_lowerL := "DB824_Error_MH_CP".Pressure[#MHConnection, #MHNumber].Warning_limit_minus,
                                 IO_Fault_Alarm_upperL := "DB824_Error_MH_CP".Pressure[#MHConnection, #MHNumber].Alarm_limit_plus,
                                 IO_Fault_Alarm_lowerL := "DB824_Error_MH_CP".Pressure[#MHConnection, #MHNumber].Alarm_limit_minus,
                                 IO_New_Fault := "DB009_Faults".Faultschanging_M1,
                                 IO_Fault_Level_1 := "DB009_Faults".Faults_FKT_Grp_1_M1,
                                 IO_Fault_Level_2 := "DB009_Faults".Faults_FKT_Grp_2_M1,
                                 IO_Fault_Level_3 := "DB009_Faults".Faults_FKT_Grp_3_M1);

           END_IF;

       END_FOR;

   END_FOR;
END_FUNCTION

FUNCTION "FC_Heating" : Void   // FC7004, SCL
{ S7_Optimized_Access := 'FALSE' }
VERSION : 0.1
   VAR_TEMP
      CompNumber : Int;
      HeatingNumber : Int;
      Real_Dummy : Real;
      TempStartTolTest : Bool;
      TempFLTGroup1 : Bool;
   END_VAR
BEGIN

   #CompNumber := 1;
   #HeatingNumber := 1;


   FOR #CompNumber := 1 TO "DB790_PlantParameter".AmountMeteringUnits DO

       FOR #HeatingNumber := 1 TO "DB753_MeteringPump".Pump[#CompNumber].AmountOfHeating DO
           #TempFLTGroup1 := 0;

           // Schritt 01: Einlesen des Prozess- Wertes
           // 
           "FC920_PV_Calc_Act_Value"(IN_Act_Value_read := "DB753_MeteringPump".Heating[#CompNumber].Exist[#HeatingNumber],
                                     IN_Act_Value_ext := FALSE,
                                     IN_Ext_Value := #Real_Dummy,
                                     IN_Read_Double := FALSE,
                                     IN_FLT_Needful := TRUE,
                                     IN_FLT_Reset := "DB009_Faults".Faults_Reset_FKT_M1,
                                     IO_Any_ArrayPV := "DB608_PV_Metering".Heating[#CompNumber].Heating[#HeatingNumber],
                                     IO_Fault_Sensor := "DB823_Error_Metering".Heating[#CompNumber].Heating[#HeatingNumber].Sensor_FLT_broken_wire,
                                     IO_New_Fault := "DB009_Faults".Faultschanging_M1,
                                     IO_FLT_Level_3 := "DB009_Faults".Faults_FKT_Grp_3_M1);

           // Schritt 02: Überwachen der Prozess- Limits
           // 
           #TempStartTolTest :=
           "DB753_MeteringPump".Heating[#CompNumber].Exist[#HeatingNumber];

           "FC916_PV_Limits"(IN_Tolerance_Test := #TempStartTolTest,
                             IN_Reset_Fault := "DB009_Faults".Faults_Reset_FKT_M1,
                             IO_Any_ArrayPV := "DB608_PV_Metering".Heating[#CompNumber].Heating[#HeatingNumber],
                             IO_Fault_Warn_upperL := "DB823_Error_Metering".Heating[#CompNumber].Heating[#HeatingNumber].Warning_limit_plus,
                             IO_Fault_Warn_lowerL := "DB823_Error_Metering".Heating[#CompNumber].Heating[#HeatingNumber].Warning_limit_minus,
                             IO_Fault_Alarm_upperL := "DB823_Error_Metering".Heating[#CompNumber].Heating[#HeatingNumber].Alarm_limit_plus,
                             IO_Fault_Alarm_lowerL := "DB823_Error_Metering".Heating[#CompNumber].Heating[#HeatingNumber].Alarm_limit_minus,
                             IO_New_Fault := "DB009_Faults".Faultschanging_M1,
                             IO_Fault_Level_1 := #TempFLTGroup1,
                             IO_Fault_Level_2 := "DB009_Faults".Faults_FKT_Grp_2_M1,
                             IO_Fault_Level_3 := "DB009_Faults".Faults_FKT_Grp_3_M1);

           "DB009_Faults".Faults_FKT_Grp_3_M1 := "DB009_Faults".Faults_FKT_Grp_3_M1 OR #TempFLTGroup1;

           // Schritt 03: Ansteuerung der Heizung
           // 
           "FC205_Tempering_1"(IN_Exist := "DB753_MeteringPump".Heating[#CompNumber].Exist[#HeatingNumber],
                               IN_Release := "DB613_Komponent_State".Heating[0].Heating[1].HeatingRelease,
                               IN_FLT_Ackn := "DB009_Faults".Faults_Reset_FKT_M1,
                               IN_actual_Temp := "DB608_PV_Metering".Heating[0].Heating[1].PV_ActV.Value,
                               IN_set_Temp := "DB608_PV_Metering".Heating[0].Heating[1].PV_SetV.Value,
                               IO_State := "DB613_Komponent_State".Heating[#CompNumber].Heating[#HeatingNumber],
                               IO_Values := "DB753_MeteringPump".HeatingController[#CompNumber].Heating[#HeatingNumber],
                               IO_Faults := "DB823_Error_Metering".Heating[#CompNumber].Heating[#HeatingNumber],
                               IO_NewFault := "DB009_Faults".Faultschanging_M1,
                               IO_FaultLevel_3 := "DB009_Faults".Faults_FKT_Grp_3_M1);


       END_FOR;

   END_FOR;
END_FUNCTION

FUNCTION "FC_ToleranceValuesComponent" : Void   // FC7006, SCL
{ S7_Optimized_Access := 'FALSE' }
VERSION : 0.1
   VAR_INPUT
      CompForShot : Array[1..16] of Bool;
      SwitchOffControl : Bool;
   END_VAR
   VAR_TEMP
      CompNumber : Int;
      TempStartTolTest : Bool;
   END_VAR
BEGIN

   #CompNumber := 1;

   FOR #CompNumber := 1 TO "DB790_PlantParameter".AmountMeteringUnits DO

       #TempStartTolTest :=
       #CompForShot[#CompNumber]
       AND "DB619_State_MPart".Cycle[1].Shotrelease
       AND NOT #SwitchOffControl;

       "FC916_PV_Limits"(IN_Tolerance_Test:=#TempStartTolTest,
                       IN_Reset_Fault:="DB009_Faults".Faults_Reset_FKT_M1,
                       IO_Any_ArrayPV:="DB608_PV_Metering".Metering[#CompNumber].Pressure,
                       IO_Fault_Warn_upperL:="DB823_Error_Metering".Pressure_Component[#CompNumber].Warning_limit_plus,
                       IO_Fault_Warn_lowerL:="DB823_Error_Metering".Pressure_Component[#CompNumber].Warning_limit_minus,
                       IO_Fault_Alarm_upperL:="DB823_Error_Metering".Pressure_Component[#CompNumber].Alarm_limit_plus,
                       IO_Fault_Alarm_lowerL:="DB823_Error_Metering".Pressure_Component[#CompNumber].Alarm_limit_minus,
                       IO_New_Fault:="DB009_Faults".Faultschanging_M1,
                       IO_Fault_Level_1:="DB009_Faults".Faults_FKT_Grp_1_M1,
                       IO_Fault_Level_2:="DB009_Faults".Faults_FKT_Grp_2_M1,
                       IO_Fault_Level_3:="DB009_Faults".Faults_FKT_Grp_3_M1);

     "FC916_PV_Limits"(IN_Tolerance_Test := #TempStartTolTest,
                       IN_Reset_Fault := "DB009_Faults".Faults_Reset_FKT_M1,
                       IO_Any_ArrayPV := "DB608_PV_Metering".Metering[#CompNumber].Flow,
                       IO_Fault_Warn_upperL := "DB823_Error_Metering".Flow_Component[#CompNumber].Warning_limit_plus,
                       IO_Fault_Warn_lowerL := "DB823_Error_Metering".Flow_Component[#CompNumber].Warning_limit_minus,
                       IO_Fault_Alarm_upperL := "DB823_Error_Metering".Flow_Component[#CompNumber].Alarm_limit_plus,
                       IO_Fault_Alarm_lowerL := "DB823_Error_Metering".Flow_Component[#CompNumber].Alarm_limit_minus,
                       IO_New_Fault := "DB009_Faults".Faultschanging_M1,
                       IO_Fault_Level_1 := "DB009_Faults".Faults_FKT_Grp_1_M1,
                       IO_Fault_Level_2 := "DB009_Faults".Faults_FKT_Grp_2_M1,
                       IO_Fault_Level_3 := "DB009_Faults".Faults_FKT_Grp_3_M1);

     "FC916_PV_Limits"(IN_Tolerance_Test := #TempStartTolTest,
                       IN_Reset_Fault := "DB009_Faults".Faults_Reset_FKT_M1,
                       IO_Any_ArrayPV := "DB608_PV_Metering".Metering[#CompNumber].MixingRatio,
                       IO_Fault_Warn_upperL := "DB823_Error_Metering".Flow_Component[#CompNumber].Warning_limit_plus_MR,
                       IO_Fault_Warn_lowerL := "DB823_Error_Metering".Flow_Component[#CompNumber].Warning_limit_minus_MR,
                       IO_Fault_Alarm_upperL := "DB823_Error_Metering".Flow_Component[#CompNumber].Alarm_limit_plus_MR,
                       IO_Fault_Alarm_lowerL := "DB823_Error_Metering".Flow_Component[#CompNumber].Alarm_limit_minus_MR,
                       IO_New_Fault := "DB009_Faults".Faultschanging_M1,
                       IO_Fault_Level_1 := "DB009_Faults".Faults_FKT_Grp_1_M1,
                       IO_Fault_Level_2 := "DB009_Faults".Faults_FKT_Grp_2_M1,
                       IO_Fault_Level_3 := "DB009_Faults".Faults_FKT_Grp_3_M1);

   END_FOR;
END_FUNCTION

FUNCTION "ShotData_01" : Void   // FC7020, SCL
{ S7_Optimized_Access := 'FALSE' }
VERSION : 0.1
   VAR_INPUT
      CompForShot : Array[1..16] of Bool;
   END_VAR
   VAR_TEMP
      MHNumber : Int;
   END_VAR
BEGIN


   #MHNumber := "DB619_State_MPart".ShotMa[1].ShotData.MH_No;

   "DB919_ShotResultMach".ShotResult_Ma[1].Component.Comp[1].ComponentActive := 0;
   "DB919_ShotResultMach".ShotResult_Ma[1].Component.Comp[2].ComponentActive := 0;
   "DB919_ShotResultMach".ShotResult_Ma[1].Component.Comp[3].ComponentActive := 0;
   "DB919_ShotResultMach".ShotResult_Ma[1].Component.Comp[4].ComponentActive := 0;
   "DB919_ShotResultMach".ShotResult_Ma[1].Component.Comp[5].ComponentActive := 0;
   "DB919_ShotResultMach".ShotResult_Ma[1].Component.Comp[6].ComponentActive := 0;


   IF "DB704_MH_Value".Mixinghead[#MHNumber].MH_Connection[1].Pump_No <> 0 THEN
       "DB919_ShotResultMach".ShotResult_Ma[1].Component.Comp[1].ComponentActive := #CompForShot["DB704_MH_Value".Mixinghead[#MHNumber].MH_Connection[1].Pump_No];
   END_IF;

   IF "DB704_MH_Value".Mixinghead[#MHNumber].MH_Connection[2].Pump_No <> 0 THEN
       "DB919_ShotResultMach".ShotResult_Ma[1].Component.Comp[2].ComponentActive := #CompForShot["DB704_MH_Value".Mixinghead[#MHNumber].MH_Connection[2].Pump_No];
   END_IF;

   IF "DB704_MH_Value".Mixinghead[#MHNumber].MH_Connection[3].Pump_No <> 0 THEN
       "DB919_ShotResultMach".ShotResult_Ma[1].Component.Comp[3].ComponentActive := #CompForShot["DB704_MH_Value".Mixinghead[#MHNumber].MH_Connection[3].Pump_No];
   END_IF;

   IF "DB704_MH_Value".Mixinghead[#MHNumber].MH_Connection[4].Pump_No <> 0 THEN
       "DB919_ShotResultMach".ShotResult_Ma[1].Component.Comp[4].ComponentActive := #CompForShot["DB704_MH_Value".Mixinghead[#MHNumber].MH_Connection[4].Pump_No];
   END_IF;

   IF "DB704_MH_Value".Mixinghead[#MHNumber].MH_Connection[5].Pump_No <> 0 THEN
       "DB919_ShotResultMach".ShotResult_Ma[1].Component.Comp[5].ComponentActive := #CompForShot["DB704_MH_Value".Mixinghead[#MHNumber].MH_Connection[5].Pump_No];
   END_IF;

   IF "DB704_MH_Value".Mixinghead[#MHNumber].MH_Connection[6].Pump_No <> 0 THEN
       "DB919_ShotResultMach".ShotResult_Ma[1].Component.Comp[6].ComponentActive := #CompForShot["DB704_MH_Value".Mixinghead[#MHNumber].MH_Connection[6].Pump_No];
   END_IF;
END_FUNCTION

FUNCTION "ShotData_OB35" : Void   // FC7021, SCL
{ S7_Optimized_Access := 'FALSE' }
VERSION : 0.1
   VAR_INPUT
      CompForShot : Array[1..16] of Bool;
   END_VAR
   VAR_TEMP
      MHNumber : Int;
      Component : Int;
      PumpNo : Int;
      Temp_CompFlowReal : Real;
      Temp_STimeReal : Real;
      TempConsumption : Real;
   END_VAR
BEGIN

   #MHNumber := "DB919_ShotResultMach".ShotResult_Ma[1].General.MH_No;

   #Temp_STimeReal := "DB606_PV_Machine".Machine[1].ShotTime.PV_ActV.Value;

   FOR #Component := 1 TO 6 DO
       #PumpNo := "DB704_MH_Value".Mixinghead[#MHNumber].MH_Connection[#Component].Pump_No;
       (* classic code: "DB919_ShotResultMach".ShotResult_Ma[1].Component.Comp[#Component].Mixingratio := 0.0;*)
       "DB919_ShotResultMach".ShotResult_Ma[1].Component.Comp[#Component].Mixingratio := REAL#0.0;
       (* classic code: "DB919_ShotResultMach".ShotResult_Ma[1].Component.Comp[#Component].Flow := 0.0;*)
       "DB919_ShotResultMach".ShotResult_Ma[1].Component.Comp[#Component].Flow := REAL#0.0;

       IF #PumpNo > 0 AND #CompForShot[#Component] = True THEN
           // Component activ? -> im FB920 ansonsten wird nach Schuss abgelöscht
           // "DB919_ShotResultMach".ShotResult_Ma[1].Component.Comp[#Component].ComponentActive := #CompForShot[#PumpNo];
           // Flow:
           #Temp_CompFlowReal := "DB919_ShotResultMach".TotalFlowShotM1[#PumpNo] / "DB919_ShotResultMach".AmountFlowValuesM1[#PumpNo];
           "DB919_ShotResultMach".ShotResult_Ma[1].Component.Comp[#Component].Flow := #Temp_CompFlowReal;
           // Ratio
           "DB919_ShotResultMach".ShotResult_Ma[1].Component.Comp[#Component].Mixingratio := "DB608_PV_Metering".Metering[#PumpNo].MixingRatio.PV_ActV.Value;
           // Consumtion
           #TempConsumption := #Temp_CompFlowReal * #Temp_STimeReal;


           IF "DB619_State_MPart".Operationmode[1].Operation AND NOT "DB619_State_MPart".ShotMa[1].ShotData.ShotDisabled THEN

